REGION Network 2: Set initial step number for the state S5
   RUNG wire#powerrail
      I_Contact( "EtatMEFhelium" )
      { S7_GenerateENO := "TRUE" } Move(in := b#0, out1 => "Data_fo_HNOSS".S5step)
   END_RUNG
   // the same network as SCL:
   IF NOT "EtatMEFhelium" THEN "Data_fo_HNOSS".S5step := b#0; END_IF;
END_REGION

REGION Network 3: Set initial step number for the state S6
   RUNG wire#powerrail
      I_Contact( "EtatMode4k" )
      { S7_GenerateENO := "TRUE" } Move(in := b#0, out1 => "Data_fo_HNOSS".S6step)
   END_RUNG
   // the same network as SCL:
   IF NOT "EtatMode4k" THEN "Data_fo_HNOSS".S6step := b#0; END_IF;
END_REGION

REGION Network 4: Set initial step number for the state S7
   RUNG wire#powerrail
      I_Contact( "EtatModeStandBy" )
      { S7_GenerateENO := "TRUE" } Move(in := b#0, out1 => "Data_fo_HNOSS".S7step)
   END_RUNG
   // the same network as SCL:
   IF NOT "EtatModeStandBy" THEN "Data_fo_HNOSS".S7step := b#0; END_IF;
END_REGION

REGION Network 5: Set initial step number for the state S8
   RUNG wire#powerrail
      I_Contact( "EtatMode2K" )
      { S7_GenerateENO := "TRUE" } Move(in := b#0, out1 => "Data_fo_HNOSS".S8step)
   END_RUNG
   // the same network as SCL:
   IF NOT "EtatMode2K" THEN "Data_fo_HNOSS".S8step := b#0; END_IF;
END_REGION

REGION Network 6: Set initial step number for the state S9 (non existent yet)
   RUNG wire#powerrail
      { S7_GenerateENO := "TRUE" } Move(in := b#0, out1 => "Data_fo_HNOSS".S9step)
   END_RUNG
   // the same network as SCL:
   "Data_fo_HNOSS".S9step := b#0;
END_REGION

REGION Network 7: Set initial step number for the state S10
   RUNG wire#powerrail
      I_Contact( "Etatrechauffage" )
      { S7_GenerateENO := "TRUE" } Move(in := b#0, out1 => "Data_fo_HNOSS".S10step)
   END_RUNG
   // the same network as SCL:
   IF NOT "Etatrechauffage" THEN "Data_fo_HNOSS".S10step := b#0; END_IF;
END_REGION

REGION Network 8: Set initial step number for the state SX (spare)
   RUNG wire#powerrail
      { S7_GenerateENO := "TRUE" } Move(in := b#0, out1 => "Data_fo_HNOSS".SXstep)
   END_RUNG
   // the same network as SCL:
   "Data_fo_HNOSS".SXstep := b#0;
END_REGION

REGION Network 9 (STL): Change to int for "compare" instruction

         L     "Data_fo_HNOSS".S4step;
         T     #S4step;
         L     "Data_fo_HNOSS".S5step;
         T     #S5step;
         L     "Data_fo_HNOSS".S6step;
         T     #S6step;
         L     "Data_fo_HNOSS".S7step;
         T     #S7step;
         L     "Data_fo_HNOSS".S8step;
         T     #S8step;
         L     "Data_fo_HNOSS".S9step;
         T     #S9step;
         L     "Data_fo_HNOSS".S10step;
         T     #S10step;
         L     "Data_fo_HNOSS".SXstep;
         T     #Sxstep;
END_REGION

REGION Network 10: Init temporary values
   RUNG wire#powerrail
      { S7_GenerateENO := "TRUE" } Move(in := 0.0, out1 => #min)
      wire#w1
      { S7_GenerateENO := "TRUE" } Move(in := 100.0, out1 => #max)
   END_RUNG
   RUNG wire#w1
      I_Contact( "Data_from_HNOSS".FV552_Closed )
      Contact( "Data_from_HNOSS".FV552_Open )
      Coil( #ToCompressor )
   END_RUNG
   // the same network as SCL:
   // ENO of a box is taken as its EN; it also drops when the box reports an error
   #min := 0.0;
   #max := 100.0;
   #ToCompressor := NOT "Data_from_HNOSS".FV552_Closed AND "Data_from_HNOSS".FV552_Open;
END_REGION

REGION Network 11: config vannes init mode
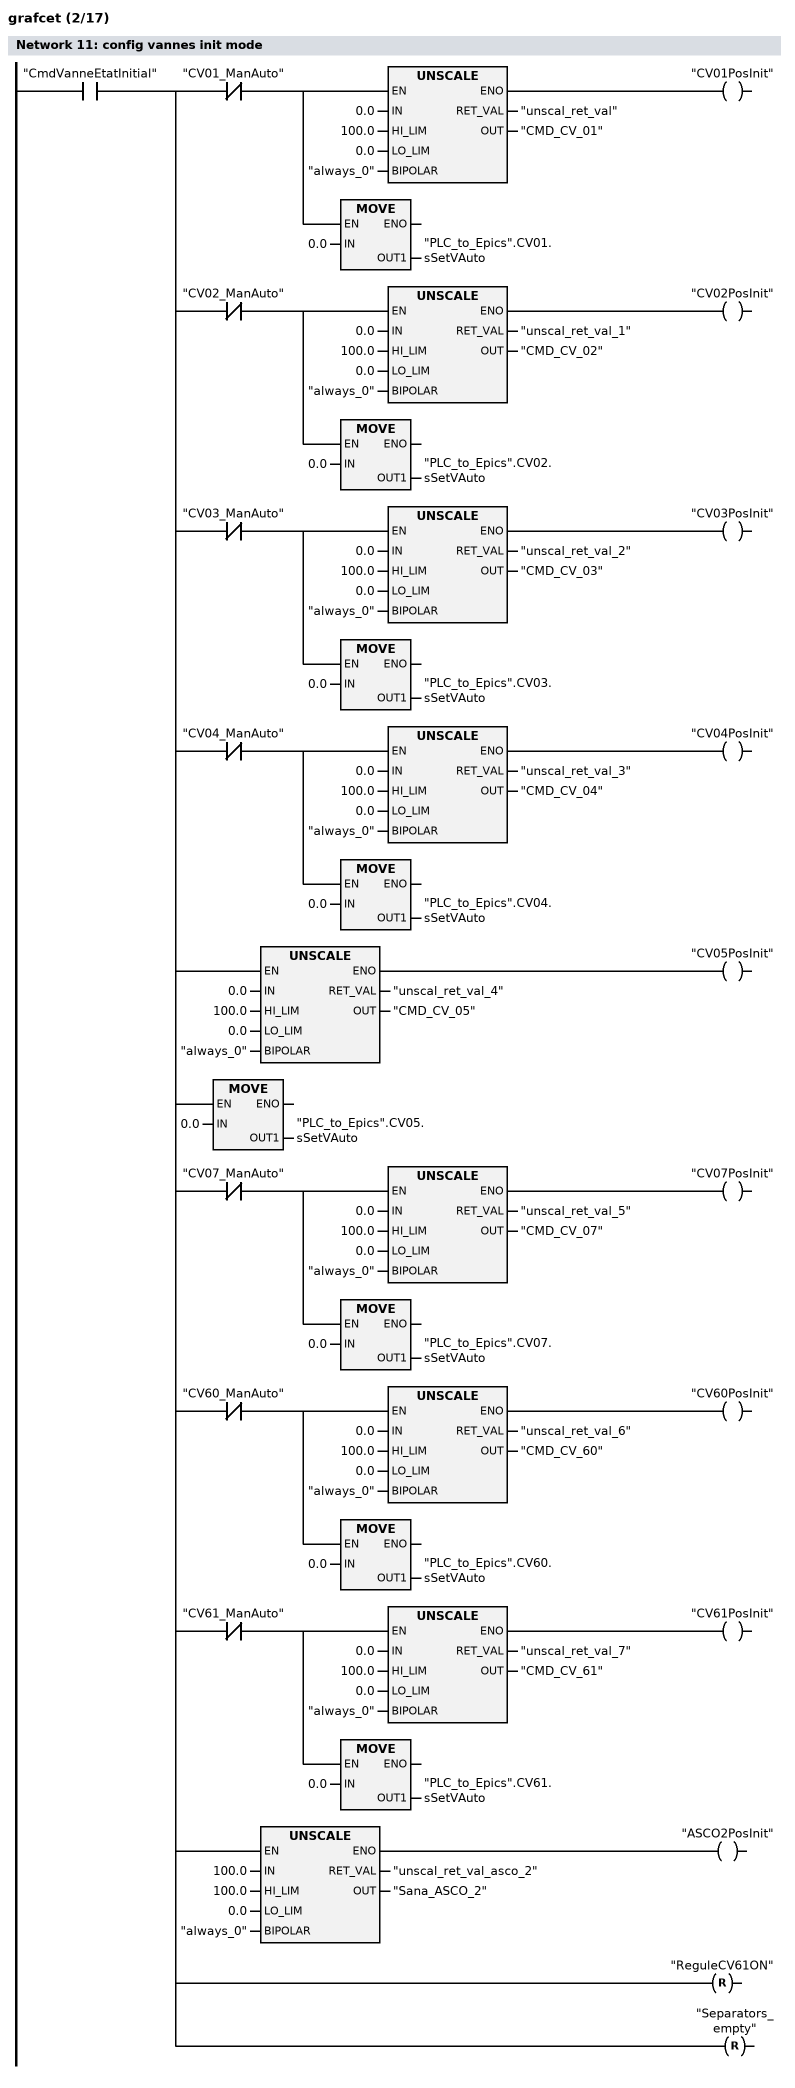
   // ENO of a box is taken as its EN; it also drops when the box reports an error
   #_w1 := "CmdVanneEtatInitial" AND NOT "CV01_ManAuto";
   #_w2 := "CmdVanneEtatInitial";
   IF #_w1 THEN
       "unscal_ret_val" := UNSCALE(in := 0.0,
                               hi_lim := 100.0,
                               lo_lim := 0.0,
                               bipolar := "always_0",
                               out => "CMD_CV_01");
   END_IF;
   "CV01PosInit" := #_w1;
   IF #_w1 THEN "PLC_to_Epics".CV01.sSetVAuto := 0.0; END_IF;
   #_w3 := #_w2 AND NOT "CV02_ManAuto";
   IF #_w3 THEN
       "unscal_ret_val_1" := UNSCALE(in := 0.0,
                               hi_lim := 100.0,
                               lo_lim := 0.0,
                               bipolar := "always_0",
                               out => "CMD_CV_02");
   END_IF;
   "CV02PosInit" := #_w3;
   IF #_w3 THEN "PLC_to_Epics".CV02.sSetVAuto := 0.0; END_IF;
   #_w4 := #_w2 AND NOT "CV03_ManAuto";
   IF #_w4 THEN
       "unscal_ret_val_2" := UNSCALE(in := 0.0,
                               hi_lim := 100.0,
                               lo_lim := 0.0,
                               bipolar := "always_0",
                               out => "CMD_CV_03");
   END_IF;
   "CV03PosInit" := #_w4;
   IF #_w4 THEN "PLC_to_Epics".CV03.sSetVAuto := 0.0; END_IF;
   #_w5 := #_w2 AND NOT "CV04_ManAuto";
   IF #_w5 THEN
       "unscal_ret_val_3" := UNSCALE(in := 0.0,
                               hi_lim := 100.0,
                               lo_lim := 0.0,
                               bipolar := "always_0",
                               out => "CMD_CV_04");
   END_IF;
   "CV04PosInit" := #_w5;
   IF #_w5 THEN "PLC_to_Epics".CV04.sSetVAuto := 0.0; END_IF;
   IF #_w2 THEN
       "unscal_ret_val_4" := UNSCALE(in := 0.0,
                               hi_lim := 100.0,
                               lo_lim := 0.0,
                               bipolar := "always_0",
                               out => "CMD_CV_05");
   END_IF;
   "CV05PosInit" := #_w2;
   IF #_w2 THEN "PLC_to_Epics".CV05.sSetVAuto := 0.0; END_IF;
   #_w6 := #_w2 AND NOT "CV07_ManAuto";
   IF #_w6 THEN
       "unscal_ret_val_5" := UNSCALE(in := 0.0,
                               hi_lim := 100.0,
                               lo_lim := 0.0,
                               bipolar := "always_0",
                               out => "CMD_CV_07");
   END_IF;
   "CV07PosInit" := #_w6;
   IF #_w6 THEN "PLC_to_Epics".CV07.sSetVAuto := 0.0; END_IF;
   #_w7 := #_w2 AND NOT "CV60_ManAuto";
   IF #_w7 THEN
       "unscal_ret_val_6" := UNSCALE(in := 0.0,
                               hi_lim := 100.0,
                               lo_lim := 0.0,
                               bipolar := "always_0",
                               out => "CMD_CV_60");
   END_IF;
   "CV60PosInit" := #_w7;
   IF #_w7 THEN "PLC_to_Epics".CV60.sSetVAuto := 0.0; END_IF;
   #_w8 := #_w2 AND NOT "CV61_ManAuto";
   IF #_w8 THEN
       "unscal_ret_val_7" := UNSCALE(in := 0.0,
                               hi_lim := 100.0,
                               lo_lim := 0.0,
                               bipolar := "always_0",
                               out => "CMD_CV_61");
   END_IF;
   "CV61PosInit" := #_w8;
   IF #_w8 THEN "PLC_to_Epics".CV61.sSetVAuto := 0.0; END_IF;
   IF #_w2 THEN
       "unscal_ret_val_asco_2" := UNSCALE(in := 100.0,
                               hi_lim := 100.0,
                               lo_lim := 0.0,
                               bipolar := "always_0",
                               out => "Sana_ASCO_2");
   END_IF;
   "ASCO2PosInit" := #_w2;
   IF #_w2 THEN
       "ReguleCV61ON" := FALSE;
       "Separators_empty" := FALSE;
   END_IF;
END_REGION

REGION Network 12: Vanne En Position Initial
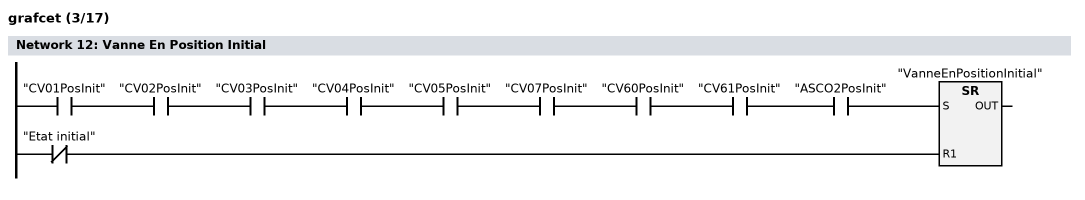
   RUNG wire#powerrail
      Contact( "CV01PosInit" )
      Contact( "CV02PosInit" )
      Contact( "CV03PosInit" )
      Contact( "CV04PosInit" )
      Contact( "CV05PosInit" )
      Contact( "CV07PosInit" )
      Contact( "CV60PosInit" )
      Contact( "CV61PosInit" )
      Contact( "ASCO2PosInit" )
      S_SR(operand := "VanneEnPositionInitial", r1 := wire#w1)
   END_RUNG
   RUNG wire#powerrail
      I_Contact( "Etat initial" )
   END_RUNG wire#w1
   // the same network as SCL:
   IF "CV01PosInit" AND "CV02PosInit" AND "CV03PosInit" AND "CV04PosInit" AND "CV05PosInit" AND "CV07PosInit" AND "CV60PosInit" AND "CV61PosInit" AND "ASCO2PosInit" THEN
       "VanneEnPositionInitial" := TRUE;   // SR flip-flop
   END_IF;
   IF NOT "Etat initial" THEN "VanneEnPositionInitial" := FALSE; END_IF;
END_REGION

REGION Network 13: config vanne etat conditionnement
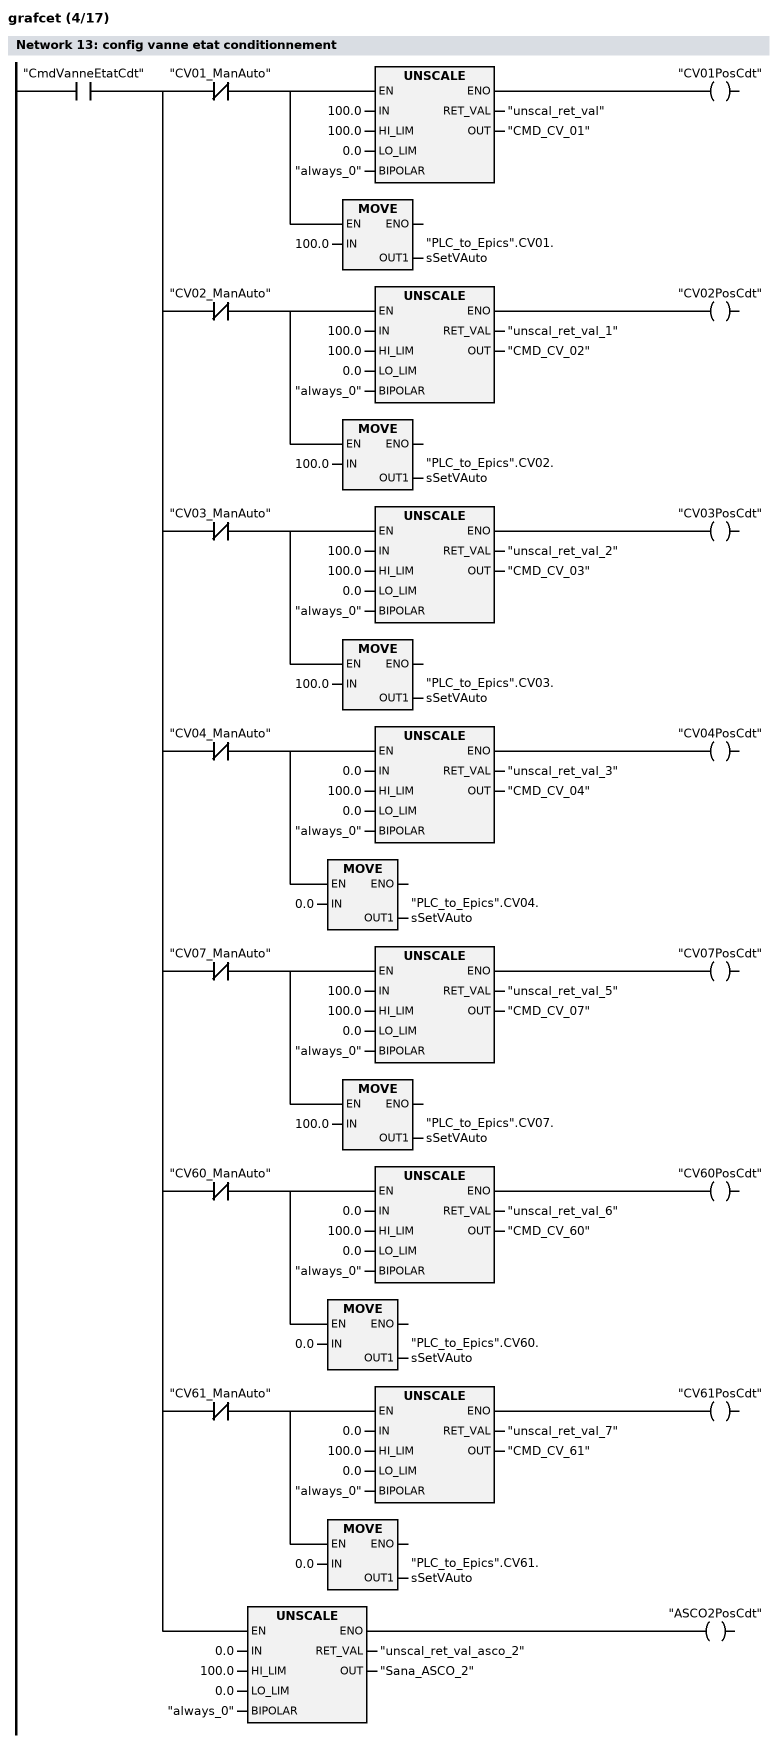
   // ENO of a box is taken as its EN; it also drops when the box reports an error
   #_w1 := "CmdVanneEtatCdt" AND NOT "CV01_ManAuto";
   #_w2 := "CmdVanneEtatCdt";
   IF #_w1 THEN
       "unscal_ret_val" := UNSCALE(in := 100.0,
                               hi_lim := 100.0,
                               lo_lim := 0.0,
                               bipolar := "always_0",
                               out => "CMD_CV_01");
   END_IF;
   "CV01PosCdt" := #_w1;
   IF #_w1 THEN "PLC_to_Epics".CV01.sSetVAuto := 100.0; END_IF;
   #_w3 := #_w2 AND NOT "CV02_ManAuto";
   IF #_w3 THEN
       "unscal_ret_val_1" := UNSCALE(in := 100.0,
                               hi_lim := 100.0,
                               lo_lim := 0.0,
                               bipolar := "always_0",
                               out => "CMD_CV_02");
   END_IF;
   "CV02PosCdt" := #_w3;
   IF #_w3 THEN "PLC_to_Epics".CV02.sSetVAuto := 100.0; END_IF;
   #_w4 := #_w2 AND NOT "CV03_ManAuto";
   IF #_w4 THEN
       "unscal_ret_val_2" := UNSCALE(in := 100.0,
                               hi_lim := 100.0,
                               lo_lim := 0.0,
                               bipolar := "always_0",
                               out => "CMD_CV_03");
   END_IF;
   "CV03PosCdt" := #_w4;
   IF #_w4 THEN "PLC_to_Epics".CV03.sSetVAuto := 100.0; END_IF;
   #_w5 := #_w2 AND NOT "CV04_ManAuto";
   IF #_w5 THEN
       "unscal_ret_val_3" := UNSCALE(in := 0.0,
                               hi_lim := 100.0,
                               lo_lim := 0.0,
                               bipolar := "always_0",
                               out => "CMD_CV_04");
   END_IF;
   "CV04PosCdt" := #_w5;
   IF #_w5 THEN "PLC_to_Epics".CV04.sSetVAuto := 0.0; END_IF;
   #_w6 := #_w2 AND NOT "CV07_ManAuto";
   IF #_w6 THEN
       "unscal_ret_val_5" := UNSCALE(in := 100.0,
                               hi_lim := 100.0,
                               lo_lim := 0.0,
                               bipolar := "always_0",
                               out => "CMD_CV_07");
   END_IF;
   "CV07PosCdt" := #_w6;
   IF #_w6 THEN "PLC_to_Epics".CV07.sSetVAuto := 100.0; END_IF;
   #_w7 := #_w2 AND NOT "CV60_ManAuto";
   IF #_w7 THEN
       "unscal_ret_val_6" := UNSCALE(in := 0.0,
                               hi_lim := 100.0,
                               lo_lim := 0.0,
                               bipolar := "always_0",
                               out => "CMD_CV_60");
   END_IF;
   "CV60PosCdt" := #_w7;
   IF #_w7 THEN "PLC_to_Epics".CV60.sSetVAuto := 0.0; END_IF;
   #_w8 := #_w2 AND NOT "CV61_ManAuto";
   IF #_w8 THEN
       "unscal_ret_val_7" := UNSCALE(in := 0.0,
                               hi_lim := 100.0,
                               lo_lim := 0.0,
                               bipolar := "always_0",
                               out => "CMD_CV_61");
   END_IF;
   "CV61PosCdt" := #_w8;
   IF #_w8 THEN "PLC_to_Epics".CV61.sSetVAuto := 0.0; END_IF;
   IF #_w2 THEN
       "unscal_ret_val_asco_2" := UNSCALE(in := 0.0,
                               hi_lim := 100.0,
                               lo_lim := 0.0,
                               bipolar := "always_0",
                               out => "Sana_ASCO_2");
   END_IF;
   "ASCO2PosCdt" := #_w2;
END_REGION

REGION Network 14: Vanne En Position Cdt
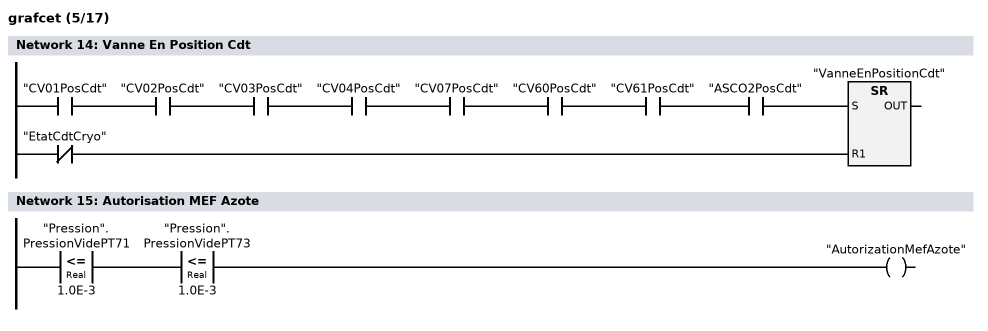
   RUNG wire#powerrail
      Contact( "CV01PosCdt" )
      Contact( "CV02PosCdt" )
      Contact( "CV03PosCdt" )
      Contact( "CV04PosCdt" )
      Contact( "CV07PosCdt" )
      Contact( "CV60PosCdt" )
      Contact( "CV61PosCdt" )
      Contact( "ASCO2PosCdt" )
      S_SR(operand := "VanneEnPositionCdt", r1 := wire#w1)
   END_RUNG
   RUNG wire#powerrail
      I_Contact( "EtatCdtCryo" )
   END_RUNG wire#w1
   // the same network as SCL:
   IF "CV01PosCdt" AND "CV02PosCdt" AND "CV03PosCdt" AND "CV04PosCdt" AND "CV07PosCdt" AND "CV60PosCdt" AND "CV61PosCdt" AND "ASCO2PosCdt" THEN
       "VanneEnPositionCdt" := TRUE;   // SR flip-flop
   END_IF;
   IF NOT "EtatCdtCryo" THEN "VanneEnPositionCdt" := FALSE; END_IF;
END_REGION

REGION Network 15: Autorisation MEF Azote
   RUNG wire#powerrail
      { S7_Templates := "SrcType := Real" } LE_Contact(in1 := "Pression".PressionVidePT71, in2 := 1.0E-3)
      { S7_Templates := "SrcType := Real" } LE_Contact(in1 := "Pression".PressionVidePT73, in2 := 1.0E-3)
      Coil( "AutorizationMefAzote" )
   END_RUNG
   // the same network as SCL:
   "AutorizationMefAzote" := ("Pression".PressionVidePT71 <= 1.0E-3) AND ("Pression".PressionVidePT73 <= 1.0E-3);
END_REGION

REGION Network 16: config vannes init mode & regule cv61 on
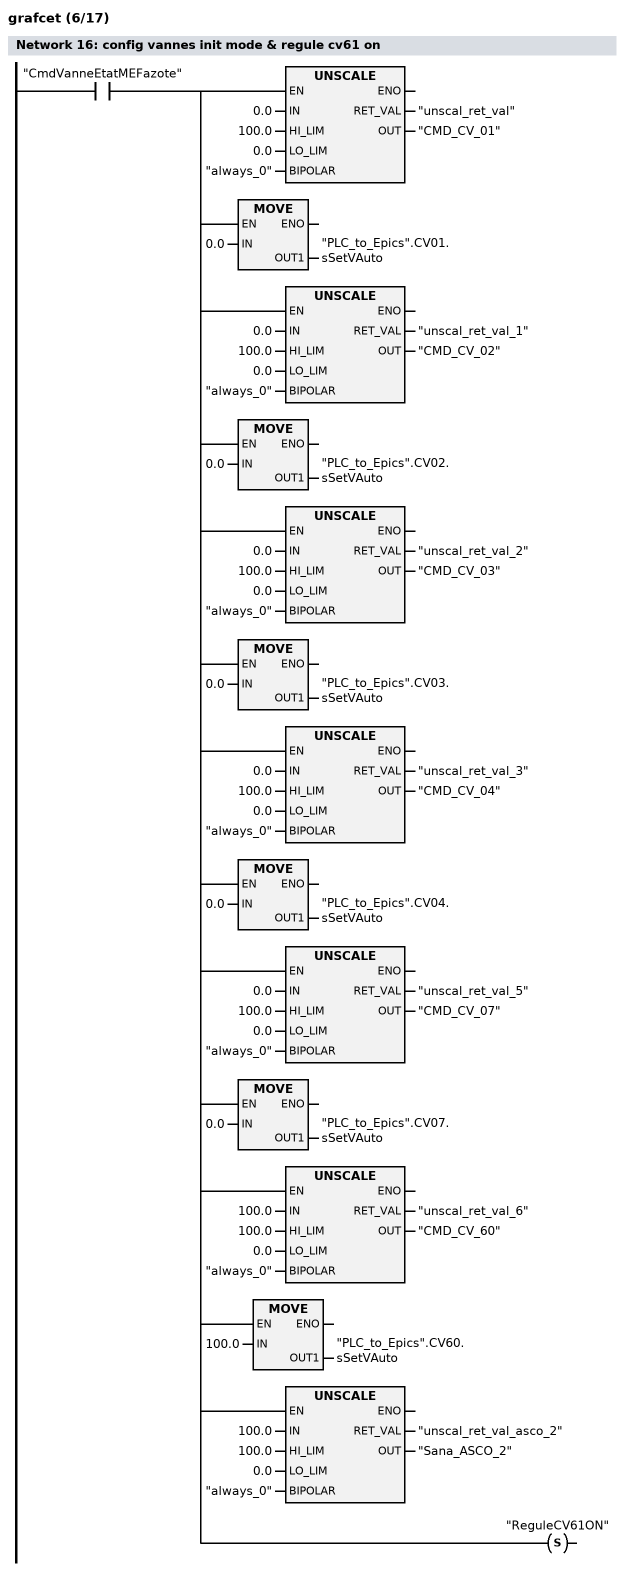
   #_w1 := "CmdVanneEtatMEFazote";
   IF #_w1 THEN
       "unscal_ret_val" := UNSCALE(in := 0.0,
                               hi_lim := 100.0,
                               lo_lim := 0.0,
                               bipolar := "always_0",
                               out => "CMD_CV_01");
       "PLC_to_Epics".CV01.sSetVAuto := 0.0;
       "unscal_ret_val_1" := UNSCALE(in := 0.0,
                               hi_lim := 100.0,
                               lo_lim := 0.0,
                               bipolar := "always_0",
                               out => "CMD_CV_02");
       "PLC_to_Epics".CV02.sSetVAuto := 0.0;
       "unscal_ret_val_2" := UNSCALE(in := 0.0,
                               hi_lim := 100.0,
                               lo_lim := 0.0,
                               bipolar := "always_0",
                               out => "CMD_CV_03");
       "PLC_to_Epics".CV03.sSetVAuto := 0.0;
       "unscal_ret_val_3" := UNSCALE(in := 0.0,
                               hi_lim := 100.0,
                               lo_lim := 0.0,
                               bipolar := "always_0",
                               out => "CMD_CV_04");
       "PLC_to_Epics".CV04.sSetVAuto := 0.0;
       "unscal_ret_val_5" := UNSCALE(in := 0.0,
                               hi_lim := 100.0,
                               lo_lim := 0.0,
                               bipolar := "always_0",
                               out => "CMD_CV_07");
       "PLC_to_Epics".CV07.sSetVAuto := 0.0;
       "unscal_ret_val_6" := UNSCALE(in := 100.0,
                               hi_lim := 100.0,
                               lo_lim := 0.0,
                               bipolar := "always_0",
                               out => "CMD_CV_60");
       "PLC_to_Epics".CV60.sSetVAuto := 100.0;
       "unscal_ret_val_asco_2" := UNSCALE(in := 100.0,
                               hi_lim := 100.0,
                               lo_lim := 0.0,
                               bipolar := "always_0",
                               out => "Sana_ASCO_2");
       "ReguleCV61ON" := TRUE;
   END_IF;
END_REGION

REGION Network 17: Régule CV61 seuil (desactive)
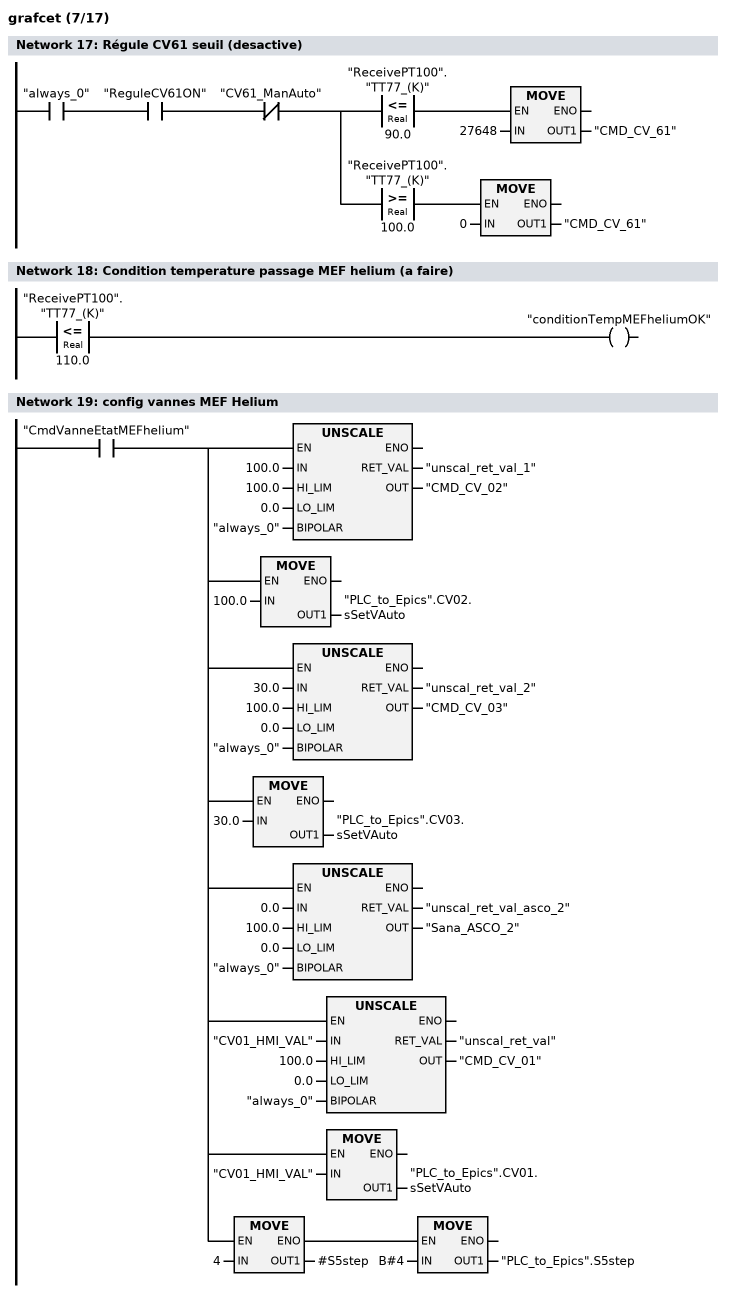
   RUNG wire#powerrail
      Contact( "always_0" )
      Contact( "ReguleCV61ON" )
      I_Contact( "CV61_ManAuto" )
      wire#w1
      { S7_Templates := "SrcType := Real" } LE_Contact(in1 := "ReceivePT100"."TT77_(K)", in2 := 90.0)
      { S7_GenerateENO := "TRUE" } Move(in := 27648, out1 => "CMD_CV_61")
   END_RUNG
   RUNG wire#w1
      { S7_Templates := "SrcType := Real" } GE_Contact(in1 := "ReceivePT100"."TT77_(K)", in2 := 100.0)
      { S7_GenerateENO := "TRUE" } Move(in := 0, out1 => "CMD_CV_61")
   END_RUNG
   // the same network as SCL:
   #_w1 := "always_0" AND "ReguleCV61ON" AND NOT "CV61_ManAuto";
   IF #_w1 AND ("ReceivePT100"."TT77_(K)" <= 90.0) THEN "CMD_CV_61" := 27648; END_IF;
   IF #_w1 AND ("ReceivePT100"."TT77_(K)" >= 100.0) THEN "CMD_CV_61" := 0; END_IF;
END_REGION

REGION Network 18: Condition temperature passage MEF helium (a faire)
   RUNG wire#powerrail
      { S7_Templates := "SrcType := Real" } LE_Contact(in1 := "ReceivePT100"."TT77_(K)", in2 := 110.0)
      Coil( "conditionTempMEFheliumOK" )
   END_RUNG
   // the same network as SCL:
   "conditionTempMEFheliumOK" := "ReceivePT100"."TT77_(K)" <= 110.0;
END_REGION

REGION Network 19: config vannes MEF Helium
   // ENO of a box is taken as its EN; it also drops when the box reports an error
   #_w1 := "CmdVanneEtatMEFhelium";
   IF #_w1 THEN
       "unscal_ret_val_1" := UNSCALE(IN := 100.0,
                               HI_LIM := 100.0,
                               LO_LIM := 0.0,
                               BIPOLAR := "always_0",
                               OUT => "CMD_CV_02");
       "PLC_to_Epics".CV02.sSetVAuto := 100.0;
       "unscal_ret_val_2" := UNSCALE(IN := 30.0,
                               HI_LIM := 100.0,
                               LO_LIM := 0.0,
                               BIPOLAR := "always_0",
                               OUT => "CMD_CV_03");
       "PLC_to_Epics".CV03.sSetVAuto := 30.0;
       "unscal_ret_val_asco_2" := UNSCALE(IN := 0.0,
                               HI_LIM := 100.0,
                               LO_LIM := 0.0,
                               BIPOLAR := "always_0",
                               OUT => "Sana_ASCO_2");
       "unscal_ret_val" := UNSCALE(IN := "CV01_HMI_VAL",
                               HI_LIM := 100.0,
                               LO_LIM := 0.0,
                               BIPOLAR := "always_0",
                               OUT => "CMD_CV_01");
       "PLC_to_Epics".CV01.sSetVAuto := "CV01_HMI_VAL";
       #S5step := 4;
       "PLC_to_Epics".S5step := B#4;
   END_IF;
END_REGION

REGION Network 20: LHe cooling down - Set step 6 (maybe setting CV03 is not needed here (done in the next network)!!!!!
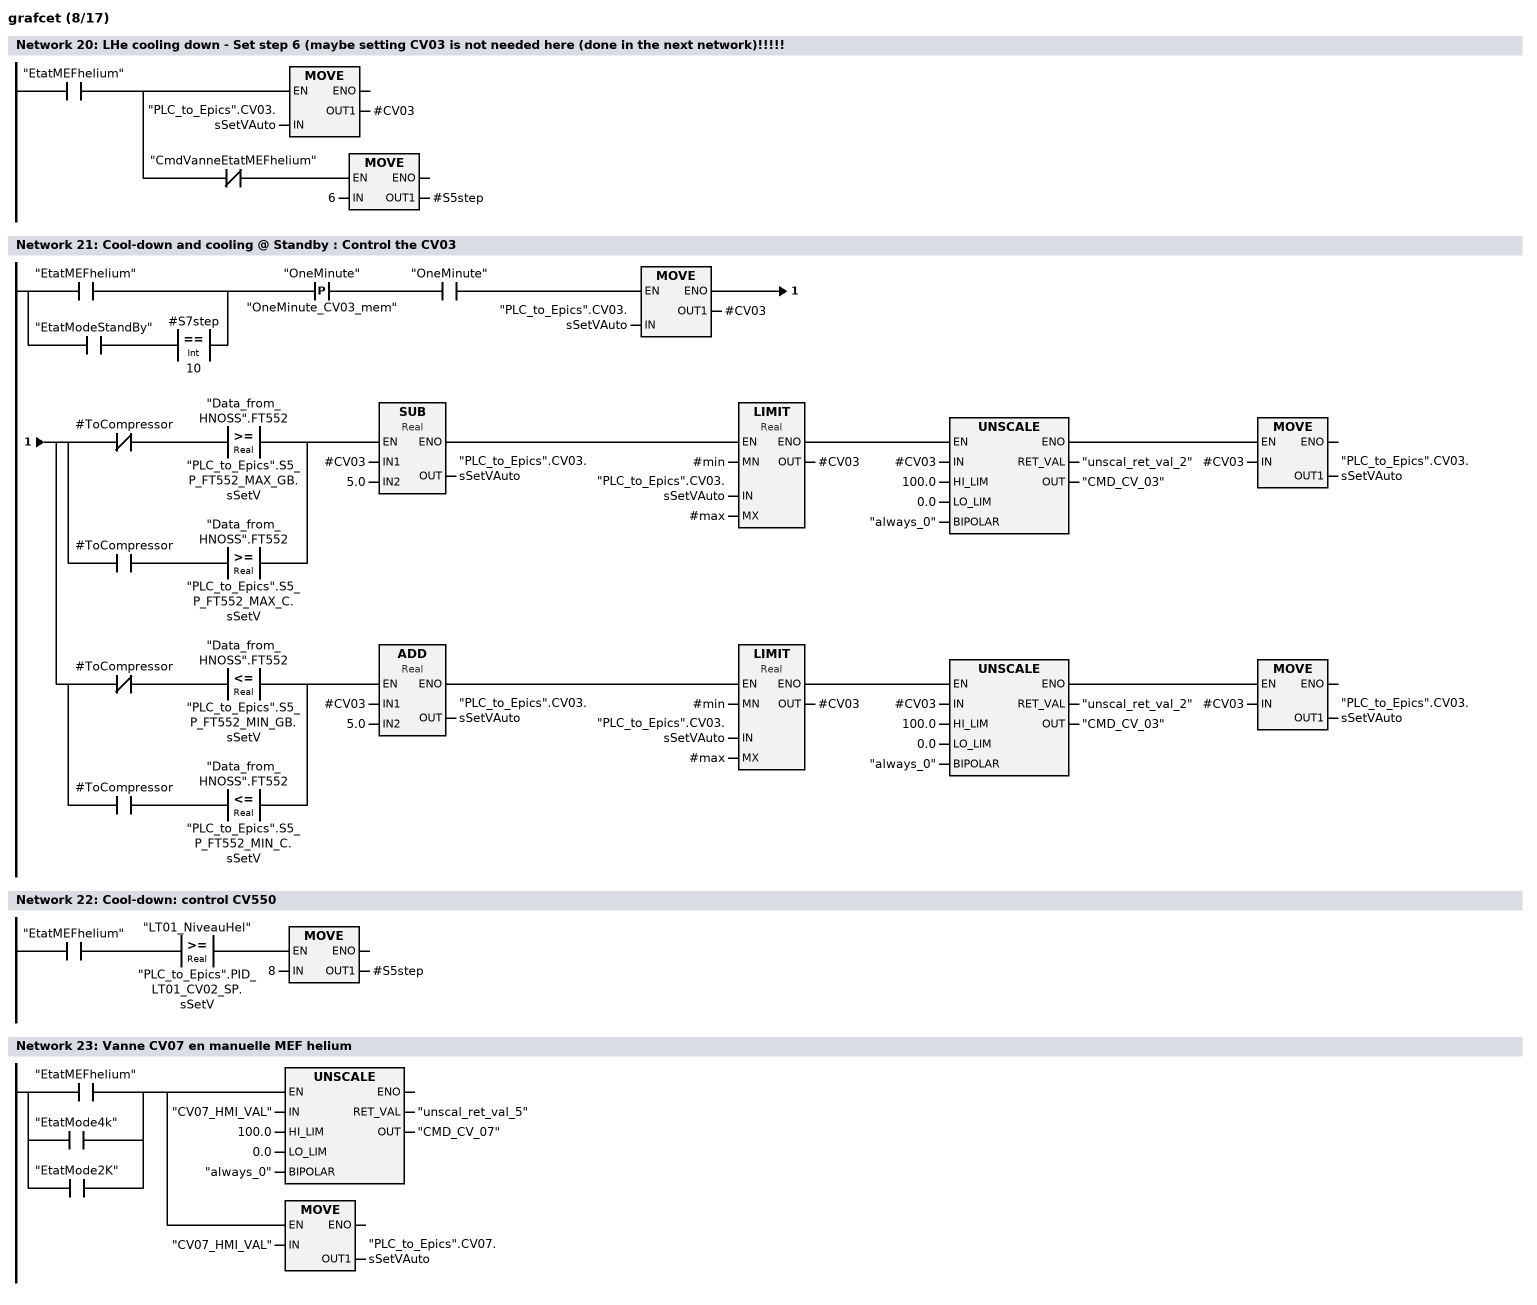
   RUNG wire#powerrail
      Contact( "EtatMEFhelium" )
      wire#w1
      { S7_GenerateENO := "TRUE" } Move(in := "PLC_to_Epics".CV03.sSetVAuto, out1 => #CV03)
   END_RUNG
   RUNG wire#w1
      I_Contact( "CmdVanneEtatMEFhelium" )
      { S7_GenerateENO := "TRUE" } Move(in := 6, out1 => #S5step)
   END_RUNG
   // the same network as SCL:
   IF "EtatMEFhelium" THEN #CV03 := "PLC_to_Epics".CV03.sSetVAuto; END_IF;
   IF "EtatMEFhelium" AND NOT "CmdVanneEtatMEFhelium" THEN #S5step := 6; END_IF;
END_REGION

REGION Network 21: Cool-down and cooling @ Standby : Control the CV03
   // ENO of a box is taken as its EN; it also drops when the box reports an error
   #_w1 := ("EtatMEFhelium" OR ("EtatModeStandBy" AND (#S7step = 10))) AND "OneMinute" AND NOT "OneMinute_CV03_mem";   // rising edge of "OneMinute"
   "OneMinute_CV03_mem" := "OneMinute";
   #_w2 := #_w1 AND "OneMinute";
   IF #_w2 THEN #CV03 := "PLC_to_Epics".CV03.sSetVAuto; END_IF;
   IF #_w2 AND ((NOT #ToCompressor AND ("Data_from_HNOSS".FT552 >= "PLC_to_Epics".S5_P_FT552_MAX_GB.sSetV)) OR (#ToCompressor AND ("Data_from_HNOSS".FT552 >= "PLC_to_Epics".S5_P_FT552_MAX_C.sSetV))) THEN
       "PLC_to_Epics".CV03.sSetVAuto := #CV03 - 5.0;
       #CV03 := LIMIT(MN := #min, IN := "PLC_to_Epics".CV03.sSetVAuto, MX := #max);
   END_IF;
   #_w3 := #_w2 AND ((NOT #ToCompressor AND ("Data_from_HNOSS".FT552 >= "PLC_to_Epics".S5_P_FT552_MAX_GB.sSetV)) OR (#ToCompressor AND ("Data_from_HNOSS".FT552 >= "PLC_to_Epics".S5_P_FT552_MAX_C.sSetV)));
   IF #_w3 THEN
       "unscal_ret_val_2" := UNSCALE(IN := #CV03,
                               HI_LIM := 100.0,
                               LO_LIM := 0.0,
                               BIPOLAR := "always_0",
                               OUT => "CMD_CV_03");
       "PLC_to_Epics".CV03.sSetVAuto := #CV03;
   END_IF;
   IF #_w2 AND ((NOT #ToCompressor AND ("Data_from_HNOSS".FT552 <= "PLC_to_Epics".S5_P_FT552_MIN_GB.sSetV)) OR (#ToCompressor AND ("Data_from_HNOSS".FT552 <= "PLC_to_Epics".S5_P_FT552_MIN_C.sSetV))) THEN
       "PLC_to_Epics".CV03.sSetVAuto := #CV03 + 5.0;
       #CV03 := LIMIT(MN := #min, IN := "PLC_to_Epics".CV03.sSetVAuto, MX := #max);
   END_IF;
   #_w4 := #_w2 AND ((NOT #ToCompressor AND ("Data_from_HNOSS".FT552 <= "PLC_to_Epics".S5_P_FT552_MIN_GB.sSetV)) OR (#ToCompressor AND ("Data_from_HNOSS".FT552 <= "PLC_to_Epics".S5_P_FT552_MIN_C.sSetV)));
   IF #_w4 THEN
       "unscal_ret_val_2" := UNSCALE(IN := #CV03,
                               HI_LIM := 100.0,
                               LO_LIM := 0.0,
                               BIPOLAR := "always_0",
                               OUT => "CMD_CV_03");
       "PLC_to_Epics".CV03.sSetVAuto := #CV03;
   END_IF;
END_REGION

REGION Network 22: Cool-down: control CV550
   RUNG wire#powerrail
      Contact( "EtatMEFhelium" )
      { S7_Templates := "SrcType := Real" } GE_Contact(in1 := "LT01_NiveauHel", in2 := "PLC_to_Epics".PID_LT01_CV02_SP.sSetV)
      { S7_GenerateENO := "TRUE" } Move(in := 8, out1 => #S5step)
   END_RUNG
   // the same network as SCL:
   IF "EtatMEFhelium" AND ("LT01_NiveauHel" >= "PLC_to_Epics".PID_LT01_CV02_SP.sSetV) THEN
       #S5step := 8;
   END_IF;
END_REGION

REGION Network 23: Vanne CV07 en manuelle MEF helium
   #_w1 := "EtatMEFhelium" OR "EtatMode4k" OR "EtatMode2K";
   IF #_w1 THEN
       "unscal_ret_val_5" := UNSCALE(in := "CV07_HMI_VAL",
                               hi_lim := 100.0,
                               lo_lim := 0.0,
                               bipolar := "always_0",
                               out => "CMD_CV_07");
       "PLC_to_Epics".CV07.sSetVAuto := "CV07_HMI_VAL";
   END_IF;
END_REGION

REGION Network 24: Vanne CV01 en manuelle MEF helium
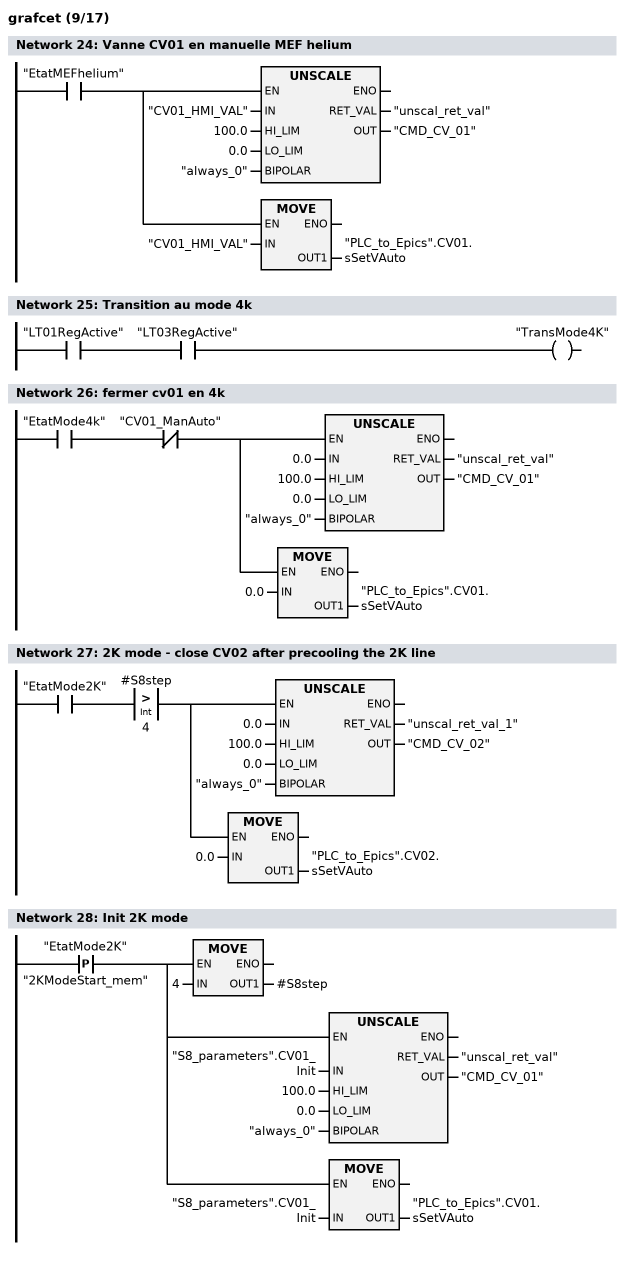
   #_w1 := "EtatMEFhelium";
   IF #_w1 THEN
       "unscal_ret_val" := UNSCALE(in := "CV01_HMI_VAL",
                               hi_lim := 100.0,
                               lo_lim := 0.0,
                               bipolar := "always_0",
                               out => "CMD_CV_01");
       "PLC_to_Epics".CV01.sSetVAuto := "CV01_HMI_VAL";
   END_IF;
END_REGION

REGION Network 25: Transition au mode 4k
   RUNG wire#powerrail
      Contact( "LT01RegActive" )
      Contact( "LT03RegActive" )
      Coil( "TransMode4K" )
   END_RUNG
   // the same network as SCL:
   "TransMode4K" := "LT01RegActive" AND "LT03RegActive";
END_REGION

REGION Network 26: fermer cv01 en 4k
   #_w1 := "EtatMode4k" AND NOT "CV01_ManAuto";
   IF #_w1 THEN
       "unscal_ret_val" := UNSCALE(in := 0.0,
                               hi_lim := 100.0,
                               lo_lim := 0.0,
                               bipolar := "always_0",
                               out => "CMD_CV_01");
       "PLC_to_Epics".CV01.sSetVAuto := 0.0;
   END_IF;
END_REGION

REGION Network 27: 2K mode - close CV02 after precooling the 2K line
   #_w1 := "EtatMode2K" AND (#S8step > 4);
   IF #_w1 THEN
       "unscal_ret_val_1" := UNSCALE(IN := 0.0,
                               HI_LIM := 100.0,
                               LO_LIM := 0.0,
                               BIPOLAR := "always_0",
                               OUT => "CMD_CV_02");
       "PLC_to_Epics".CV02.sSetVAuto := 0.0;
   END_IF;
END_REGION

REGION Network 28: Init 2K mode
   #_w1 := "EtatMode2K" AND NOT "2KModeStart_mem";   // rising edge of "EtatMode2K"
   "2KModeStart_mem" := "EtatMode2K";
   IF #_w1 THEN
       #S8step := 4;
       "unscal_ret_val" := UNSCALE(IN := "S8_parameters".CV01_Init,
                               HI_LIM := 100.0,
                               LO_LIM := 0.0,
                               BIPOLAR := "always_0",
                               OUT => "CMD_CV_01");
       "PLC_to_Epics".CV01.sSetVAuto := "S8_parameters".CV01_Init;
   END_IF;
END_REGION

REGION Network 29: 2K mode - precooling (step4)
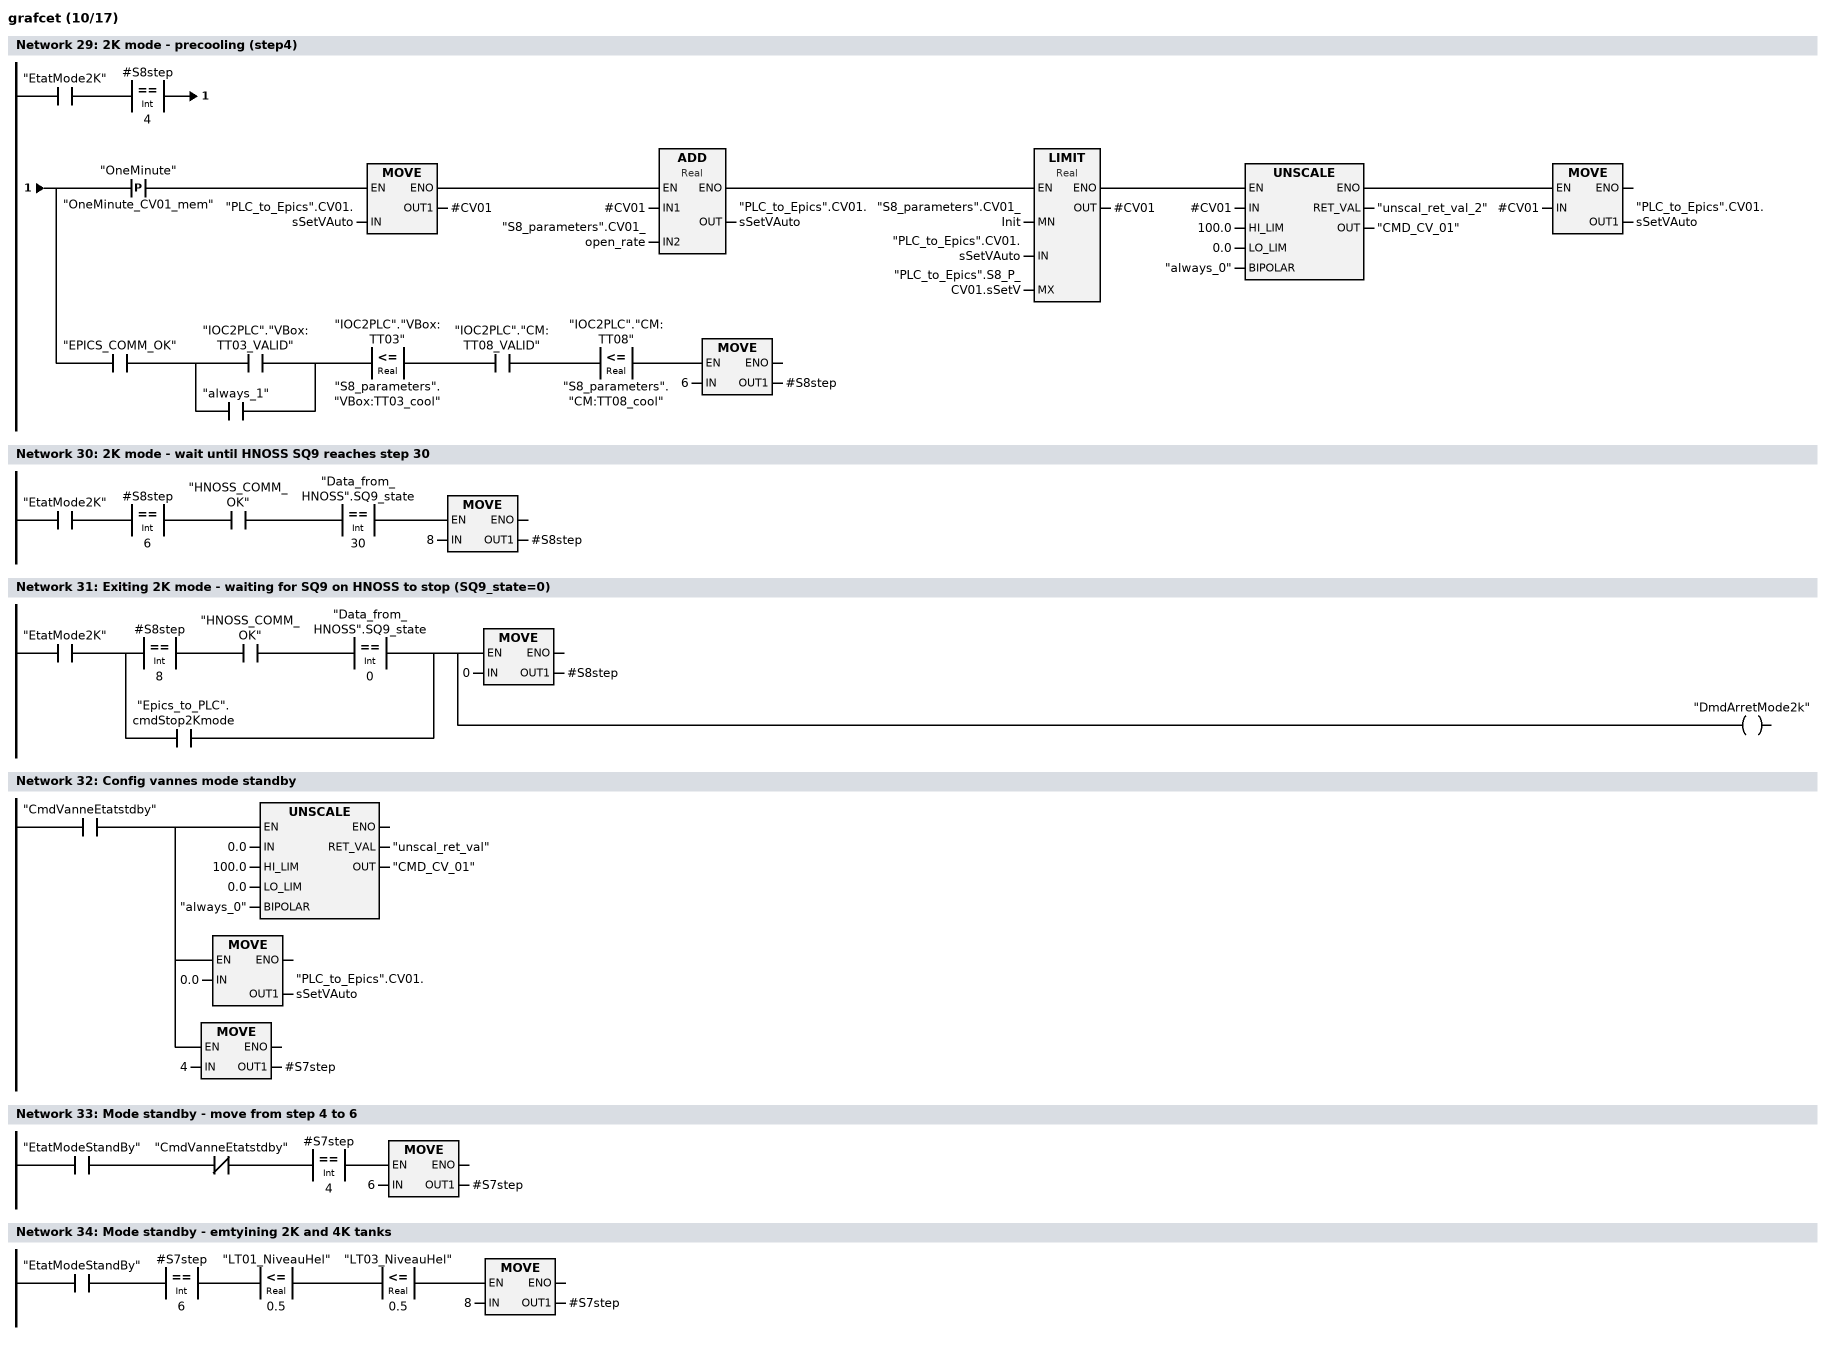
   // ENO of a box is taken as its EN; it also drops when the box reports an error
   #_w1 := "EtatMode2K" AND (#S8step = 4);
   #_w2 := #_w1 AND "OneMinute" AND NOT "OneMinute_CV01_mem";   // rising edge of "OneMinute"
   "OneMinute_CV01_mem" := "OneMinute";
   IF #_w2 THEN
       #CV01 := "PLC_to_Epics".CV01.sSetVAuto;
       "PLC_to_Epics".CV01.sSetVAuto := #CV01 + "S8_parameters".CV01_open_rate;
       #CV01 := LIMIT(MN := "S8_parameters".CV01_Init, IN := "PLC_to_Epics".CV01.sSetVAuto, MX := "PLC_to_Epics".S8_P_CV01.sSetV);